VERSION : 0.1
BEGIN

REGION Network 1
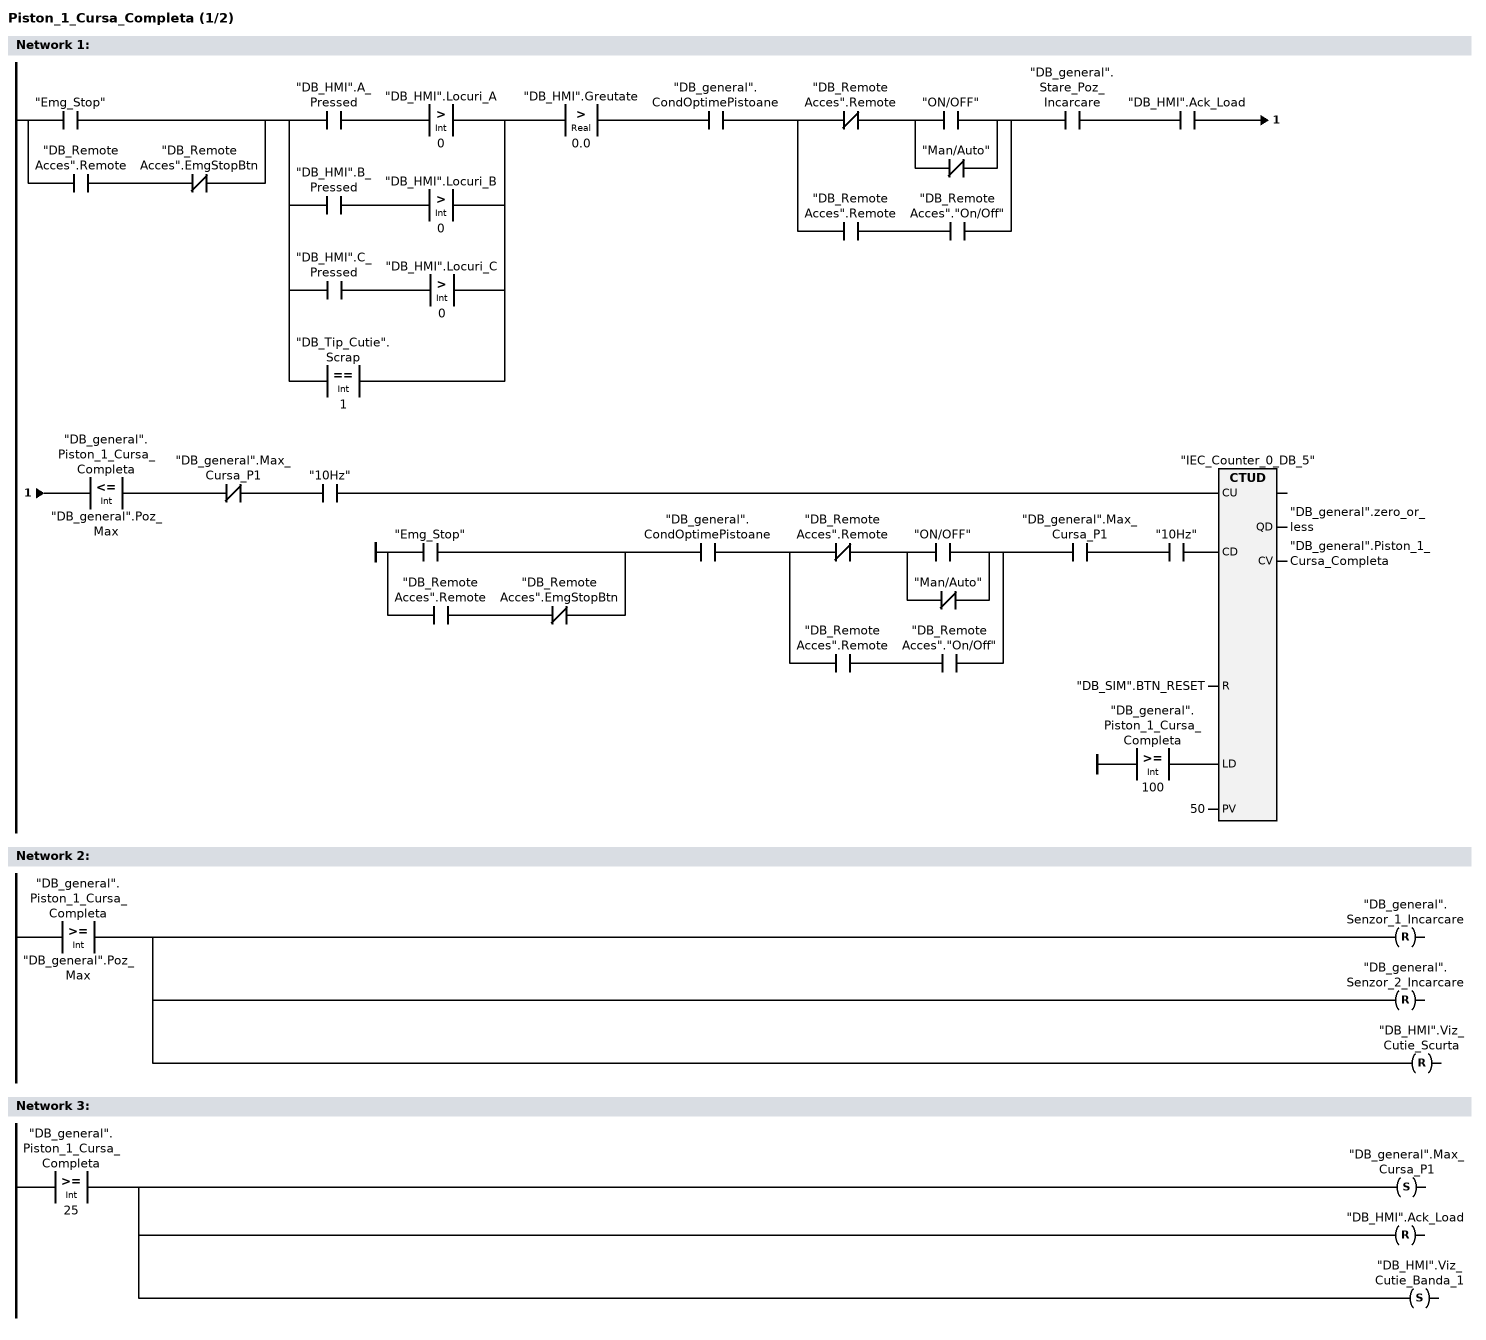
   "IEC_Counter_0_DB_5".CTUD(CU := ("Emg_Stop" OR ("DB_RemoteAcces".Remote AND NOT "DB_RemoteAcces".EmgStopBtn)) AND (("DB_HMI".A_Pressed AND ("DB_HMI".Locuri_A > 0)) OR ("DB_HMI".B_Pressed AND ("DB_HMI".Locuri_B > 0)) OR ("DB_HMI".C_Pressed AND ("DB_HMI".Locuri_C > 0)) OR ("DB_Tip_Cutie".Scrap = 1)) AND ("DB_HMI".Greutate > 0.0) AND "DB_general".CondOptimePistoane AND ((NOT "DB_RemoteAcces".Remote AND ("ON/OFF" OR NOT "Man/Auto")) OR ("DB_RemoteAcces".Remote AND "DB_RemoteAcces"."On/Off")) AND "DB_general".Stare_Poz_Incarcare AND "DB_HMI".Ack_Load AND ("DB_general".Piston_1_Cursa_Completa <= "DB_general".Poz_Max) AND NOT "DB_general".Max_Cursa_P1 AND "10Hz",
                           CD := ("Emg_Stop" OR ("DB_RemoteAcces".Remote AND NOT "DB_RemoteAcces".EmgStopBtn)) AND "DB_general".CondOptimePistoane AND ((NOT "DB_RemoteAcces".Remote AND ("ON/OFF" OR NOT "Man/Auto")) OR ("DB_RemoteAcces".Remote AND "DB_RemoteAcces"."On/Off")) AND "DB_general".Max_Cursa_P1 AND "10Hz",
                           R := "DB_SIM".BTN_RESET,
                           LD := "DB_general".Piston_1_Cursa_Completa >= 100,
                           PV := 50,
                           QD => "DB_general".zero_or_less,
                           CV => "DB_general".Piston_1_Cursa_Completa);
END_REGION

REGION Network 2
   RUNG wire#powerrail
      { S7_Templates := "SrcType := Int" } GE_Contact(in1 := "DB_general".Piston_1_Cursa_Completa, in2 := "DB_general".Poz_Max)
      wire#w1
      R_Coil( "DB_general".Senzor_1_Incarcare )
   END_RUNG
   RUNG wire#w1
      R_Coil( "DB_general".Senzor_2_Incarcare )
   END_RUNG
   RUNG wire#w1
      R_Coil( "DB_HMI".Viz_Cutie_Scurta )
   END_RUNG
   // the same network as SCL:
   IF "DB_general".Piston_1_Cursa_Completa >= "DB_general".Poz_Max THEN
       "DB_general".Senzor_1_Incarcare := FALSE;
       "DB_general".Senzor_2_Incarcare := FALSE;
       "DB_HMI".Viz_Cutie_Scurta := FALSE;
   END_IF;
END_REGION

REGION Network 3
   RUNG wire#powerrail
      { S7_Templates := "SrcType := Int" } GE_Contact(in1 := "DB_general".Piston_1_Cursa_Completa, in2 := 25)
      wire#w1
      S_Coil( "DB_general".Max_Cursa_P1 )
   END_RUNG
   RUNG wire#w1
      R_Coil( "DB_HMI".Ack_Load )
   END_RUNG
   RUNG wire#w1
      S_Coil( "DB_HMI".Viz_Cutie_Banda_1 )
   END_RUNG
   // the same network as SCL:
   IF "DB_general".Piston_1_Cursa_Completa >= 25 THEN
       "DB_general".Max_Cursa_P1 := TRUE;
       "DB_HMI".Ack_Load := FALSE;
       "DB_HMI".Viz_Cutie_Banda_1 := TRUE;
   END_IF;
END_REGION

REGION Network 4
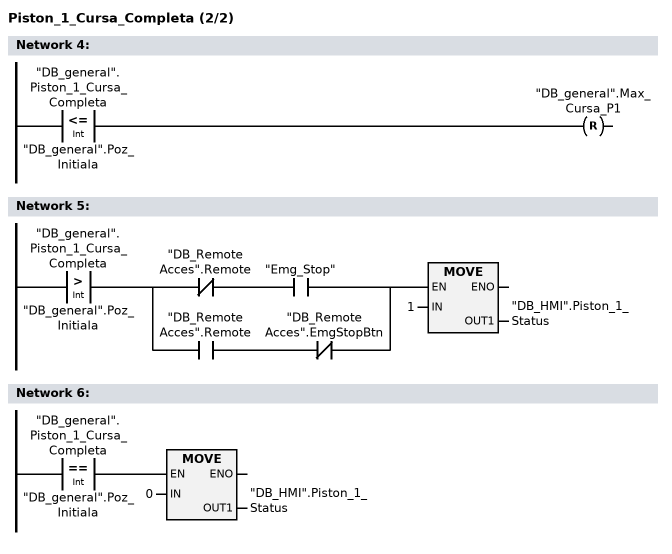
   RUNG wire#powerrail
      { S7_Templates := "SrcType := Int" } LE_Contact(in1 := "DB_general".Piston_1_Cursa_Completa, in2 := "DB_general".Poz_Initiala)
      R_Coil( "DB_general".Max_Cursa_P1 )
   END_RUNG
   // the same network as SCL:
   IF "DB_general".Piston_1_Cursa_Completa <= "DB_general".Poz_Initiala THEN
       "DB_general".Max_Cursa_P1 := FALSE;
   END_IF;
END_REGION

REGION Network 5
   RUNG wire#powerrail
      { S7_Templates := "SrcType := Int" } GT_Contact(in1 := "DB_general".Piston_1_Cursa_Completa, in2 := "DB_general".Poz_Initiala)
      wire#w1
      I_Contact( "DB_RemoteAcces".Remote )
      Contact( "Emg_Stop" )
      wire#w2
      { S7_GenerateENO := "TRUE" } Move(in := 1, out1 => "DB_HMI".Piston_1_Status)
   END_RUNG
   RUNG wire#w1
      Contact( "DB_RemoteAcces".Remote )
      I_Contact( "DB_RemoteAcces".EmgStopBtn )
   END_RUNG wire#w2
   // the same network as SCL:
   IF ("DB_general".Piston_1_Cursa_Completa > "DB_general".Poz_Initiala) AND ((NOT "DB_RemoteAcces".Remote AND "Emg_Stop") OR ("DB_RemoteAcces".Remote AND NOT "DB_RemoteAcces".EmgStopBtn)) THEN
       "DB_HMI".Piston_1_Status := 1;
   END_IF;
END_REGION

REGION Network 6
   RUNG wire#powerrail
      { S7_Templates := "SrcType := Int" } EQ_Contact(in1 := "DB_general".Piston_1_Cursa_Completa, in2 := "DB_general".Poz_Initiala)
      { S7_GenerateENO := "TRUE" } Move(in := 0, out1 => "DB_HMI".Piston_1_Status)
   END_RUNG
   // the same network as SCL:
   IF "DB_general".Piston_1_Cursa_Completa = "DB_general".Poz_Initiala THEN
       "DB_HMI".Piston_1_Status := 0;
   END_IF;
END_REGION
END_FUNCTION_BLOCK

FUNCTION_BLOCK "Piston_2_Cursa_Completa"   // FB17, LAD
{ S7_Optimized_Access := 'FALSE' }
VERSION : 0.1
BEGIN

REGION Network 1
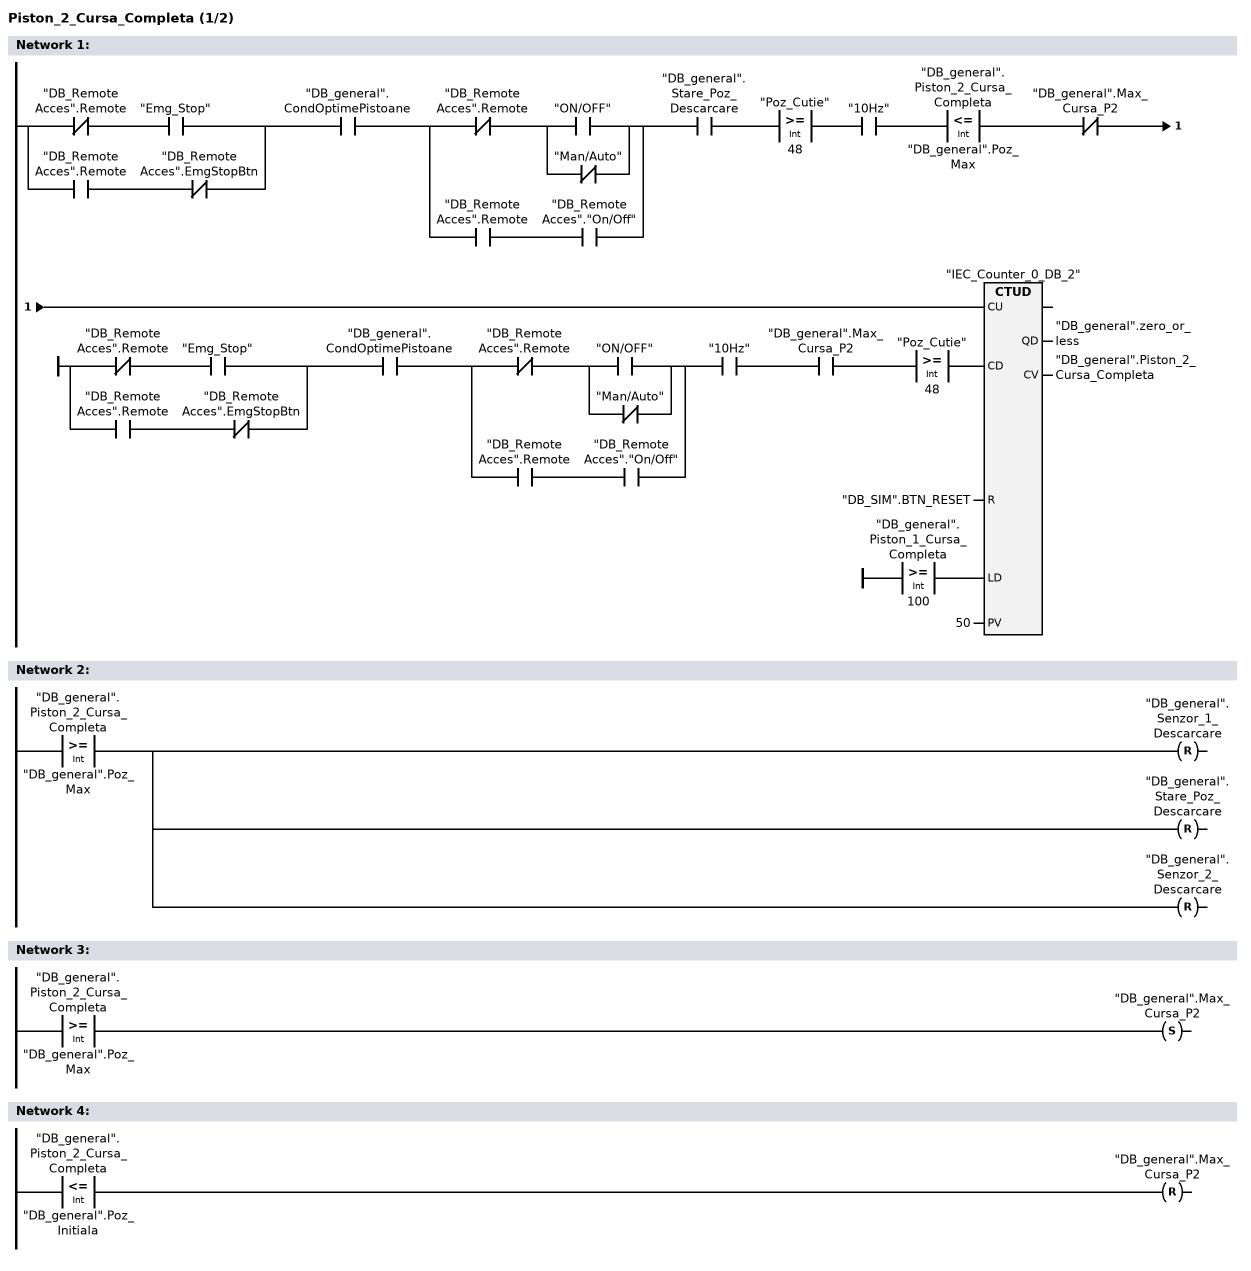
   "IEC_Counter_0_DB_2".CTUD(CU := ((NOT "DB_RemoteAcces".Remote AND "Emg_Stop") OR ("DB_RemoteAcces".Remote AND NOT "DB_RemoteAcces".EmgStopBtn)) AND "DB_general".CondOptimePistoane AND ((NOT "DB_RemoteAcces".Remote AND ("ON/OFF" OR NOT "Man/Auto")) OR ("DB_RemoteAcces".Remote AND "DB_RemoteAcces"."On/Off")) AND "DB_general".Stare_Poz_Descarcare AND ("Poz_Cutie" >= 48) AND "10Hz" AND ("DB_general".Piston_2_Cursa_Completa <= "DB_general".Poz_Max) AND NOT "DB_general".Max_Cursa_P2,
                           CD := ((NOT "DB_RemoteAcces".Remote AND "Emg_Stop") OR ("DB_RemoteAcces".Remote AND NOT "DB_RemoteAcces".EmgStopBtn)) AND "DB_general".CondOptimePistoane AND ((NOT "DB_RemoteAcces".Remote AND ("ON/OFF" OR NOT "Man/Auto")) OR ("DB_RemoteAcces".Remote AND "DB_RemoteAcces"."On/Off")) AND "10Hz" AND "DB_general".Max_Cursa_P2 AND ("Poz_Cutie" >= 48),
                           R := "DB_SIM".BTN_RESET,
                           LD := "DB_general".Piston_1_Cursa_Completa >= 100,
                           PV := 50,
                           QD => "DB_general".zero_or_less,
                           CV => "DB_general".Piston_2_Cursa_Completa);
END_REGION

REGION Network 2
   RUNG wire#powerrail
      { S7_Templates := "SrcType := Int" } GE_Contact(in1 := "DB_general".Piston_2_Cursa_Completa, in2 := "DB_general".Poz_Max)
      wire#w1
      R_Coil( "DB_general".Senzor_1_Descarcare )
   END_RUNG
   RUNG wire#w1
      R_Coil( "DB_general".Stare_Poz_Descarcare )
   END_RUNG
   RUNG wire#w1
      R_Coil( "DB_general".Senzor_2_Descarcare )
   END_RUNG
   // the same network as SCL:
   IF "DB_general".Piston_2_Cursa_Completa >= "DB_general".Poz_Max THEN
       "DB_general".Senzor_1_Descarcare := FALSE;
       "DB_general".Stare_Poz_Descarcare := FALSE;
       "DB_general".Senzor_2_Descarcare := FALSE;
   END_IF;
END_REGION

REGION Network 3
   RUNG wire#powerrail
      { S7_Templates := "SrcType := Int" } GE_Contact(in1 := "DB_general".Piston_2_Cursa_Completa, in2 := "DB_general".Poz_Max)
      S_Coil( "DB_general".Max_Cursa_P2 )
   END_RUNG
   // the same network as SCL:
   IF "DB_general".Piston_2_Cursa_Completa >= "DB_general".Poz_Max THEN
       "DB_general".Max_Cursa_P2 := TRUE;
   END_IF;
END_REGION

REGION Network 4
   RUNG wire#powerrail
      { S7_Templates := "SrcType := Int" } LE_Contact(in1 := "DB_general".Piston_2_Cursa_Completa, in2 := "DB_general".Poz_Initiala)
      R_Coil( "DB_general".Max_Cursa_P2 )
   END_RUNG
   // the same network as SCL:
   IF "DB_general".Piston_2_Cursa_Completa <= "DB_general".Poz_Initiala THEN
       "DB_general".Max_Cursa_P2 := FALSE;
   END_IF;
END_REGION

REGION Network 5
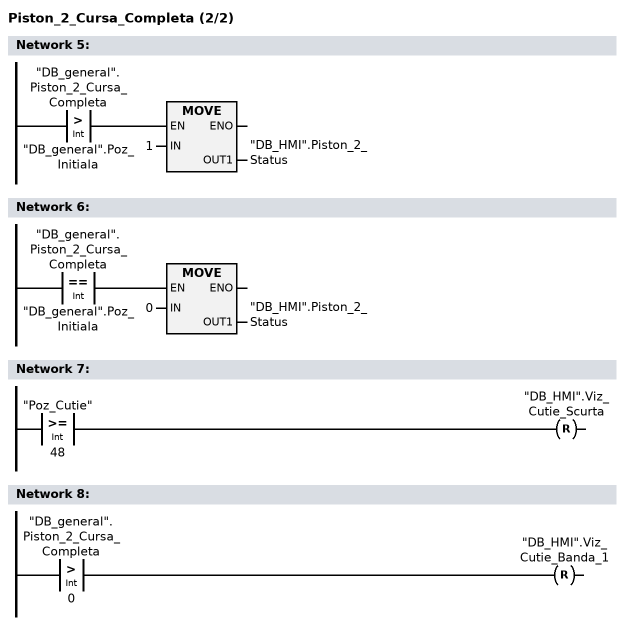
   RUNG wire#powerrail
      { S7_Templates := "SrcType := Int" } GT_Contact(in1 := "DB_general".Piston_2_Cursa_Completa, in2 := "DB_general".Poz_Initiala)
      { S7_GenerateENO := "TRUE" } Move(in := 1, out1 => "DB_HMI".Piston_2_Status)
   END_RUNG
   // the same network as SCL:
   IF "DB_general".Piston_2_Cursa_Completa > "DB_general".Poz_Initiala THEN
       "DB_HMI".Piston_2_Status := 1;
   END_IF;
END_REGION

REGION Network 6
   RUNG wire#powerrail
      { S7_Templates := "SrcType := Int" } EQ_Contact(in1 := "DB_general".Piston_2_Cursa_Completa, in2 := "DB_general".Poz_Initiala)
      { S7_GenerateENO := "TRUE" } Move(in := 0, out1 => "DB_HMI".Piston_2_Status)
   END_RUNG
   // the same network as SCL:
   IF "DB_general".Piston_2_Cursa_Completa = "DB_general".Poz_Initiala THEN
       "DB_HMI".Piston_2_Status := 0;
   END_IF;
END_REGION

REGION Network 7
   RUNG wire#powerrail
      { S7_Templates := "SrcType := Int" } GE_Contact(in1 := "Poz_Cutie", in2 := 48)
      R_Coil( "DB_HMI".Viz_Cutie_Scurta )
   END_RUNG
   // the same network as SCL:
   IF "Poz_Cutie" >= 48 THEN "DB_HMI".Viz_Cutie_Scurta := FALSE; END_IF;
END_REGION

REGION Network 8
   RUNG wire#powerrail
      { S7_Templates := "SrcType := Int" } GT_Contact(in1 := "DB_general".Piston_2_Cursa_Completa, in2 := 0)
      R_Coil( "DB_HMI".Viz_Cutie_Banda_1 )
   END_RUNG
   // the same network as SCL:
   IF "DB_general".Piston_2_Cursa_Completa > 0 THEN "DB_HMI".Viz_Cutie_Banda_1 := FALSE; END_IF;
END_REGION
END_FUNCTION_BLOCK

// folder: Statie Distribuire/Functii

FUNCTION_BLOCK "Banda_1"   // FB4, SCL
{ S7_Optimized_Access := 'FALSE' }
VERSION : 0.1
   VAR_INPUT
      Stare_Poz_Incarcare : Bool;
      Stare_Poz_Descarcare : Bool;
      Stare_Descarcare : Bool;   // Acesta este o valoare de test in care urm ca la finalul de cursa (Animatie Banda 1) pozitia descarcare sa fie facuta adev
      "Man/Auto" : Bool;
      Btn_LOAD : Bool;
   END_VAR
   VAR_OUTPUT
      Status_Banda_1 : Bool;
   END_VAR
   VAR
      Status_Poz_Cantar : Bool;
      Greutate_cantar : Int;
      Limitare_Interval : Bool;
      "ON/OFF" : Bool;
      Start_Pressed : Bool;
      AFost : Bool;
      Aux : Bool;
      LOAD_Pressed : Bool;
   END_VAR
BEGIN
   //MOD MANUAL/AUTOMAT + BUTOANE MANUAL
   IF #"Man/Auto"  THEN//daca e modul manual poti actiona butoane  true e manual false e automat

       IF "Start"  THEN
           #"Start_Pressed" := TRUE;  // setare variabila aux
           #"ON/OFF" := #Start_Pressed;
           "ON/OFF" := #"ON/OFF";
       END_IF;

       IF  "Stop"=TRUE  THEN
           #"ON/OFF" := #Start_Pressed;  //atribuire var aux
           "ON/OFF" := #"ON/OFF";
       ELSE
           IF "Stop" = FALSE THEN
               #"ON/OFF" := FALSE;
               "ON/OFF" := #"ON/OFF";
               #"Start_Pressed" := FALSE;
           END_IF;// reset variabila auxiliară la apasare stop
       END_IF;
       IF "Emg_Stop" = TRUE  THEN
           #"ON/OFF" := #Start_Pressed;  //atribuire var aux
       ELSE
           IF "Emg_Stop" = FALSE  THEN
               #"ON/OFF" := FALSE;
               "ON/OFF" := #"ON/OFF";
               #"Start_Pressed" := FALSE;
           END_IF;// reset variabila auxiliară la apasare stop
       END_IF;


   ELSE
      // #"ON/OFF" := FALSE;
      // "ON/OFF" := #"ON/OFF";
      #"Start_Pressed" := FALSE;  // Resetați variabila auxiliară în modul Manual


   END_IF;


   //LIMITARI CAPAT DE BANDA

   IF #Stare_Poz_Incarcare AND #Stare_Poz_Descarcare = FALSE AND #Stare_Descarcare=FALSE THEN//limitari de la sezorii din capetele benzii
       #Limitare_Interval := FALSE; //daca e prezent la primul nu porneste 
   ELSE
       IF #Stare_Poz_Incarcare = FALSE AND #Stare_Poz_Descarcare AND #Stare_Descarcare THEN
         #Limitare_Interval := FALSE;//daca e prezent la al doilea se opreste banda
     ELSE
         #Limitare_Interval := TRUE;

     END_IF;


   END_IF;
   // Logica pentru setare și resetare


   //START MOTOARE 
   IF #Btn_LOAD THEN
       #LOAD_Pressed := true;
   END_IF;

   IF "Poz_Cutie"<=100 THEN

       #LOAD_Pressed := TRUE;

   ELSE
       #LOAD_Pressed := FALSE;
       // Statement section IF
       ;
   END_IF;

   IF "DB_RemoteAcces"."Remote" = FALSE THEN

       IF "Man/Auto" THEN
           IF "Emg_Stop" = TRUE AND #"ON/OFF" = TRUE AND #Limitare_Interval AND "DB_HMI".BTN_LOAD THEN


               #Status_Banda_1 := TRUE;

           ELSE

               #Status_Banda_1 := FALSE;
           END_IF;

       ELSE
           IF "Emg_Stop" = TRUE AND #Limitare_Interval AND "DB_HMI".BTN_LOAD THEN

               #Status_Banda_1 := TRUE;
           ELSE

               #Status_Banda_1 := FALSE;
           END_IF;


       END_IF;


   ELSE
       IF "DB_RemoteAcces"."Remote" = TRUE THEN
           IF "DB_RemoteAcces"."Manual/Auto" = FALSE THEN
               IF "DB_RemoteAcces".EmgStopBtn = FALSE AND "DB_RemoteAcces"."On/Off" = TRUE AND #Limitare_Interval AND "DB_HMI".BTN_LOAD THEN


                   #Status_Banda_1 := TRUE;

               ELSE

                   #Status_Banda_1 := FALSE;
               END_IF;

           ELSE
               IF "DB_RemoteAcces".EmgStopBtn= FALSE AND "DB_RemoteAcces"."On/Off" = TRUE AND #Limitare_Interval AND"DB_HMI".BTN_LOAD THEN

                   #Status_Banda_1 := TRUE;
               ELSE

                   #Status_Banda_1 := FALSE;
               END_IF;


           END_IF;
       END_IF;

   END_IF;
END_FUNCTION_BLOCK

FUNCTION_BLOCK "Cantar"   // FB6, SCL
{ S7_Optimized_Access := 'FALSE' }
VERSION : 0.1
   VAR_INPUT
      Status_Poz : Bool;
      emgy_ok : Bool;
   END_VAR
   VAR_OUTPUT
      Greutate : Int;
   END_VAR
   VAR
      time_struct : Struct
         an : Byte;
         luna : Byte;
         zi : Byte;
         ora : Byte;
         minut : Byte;
         sec : Byte;
         milisec : Byte;
         weekday : Byte;
      END_STRUCT;
      rand : Int;
      i : Int;
      val : Int := 100;
   END_VAR
BEGIN

   #val := 100;

   IF "Emg_Stop" = TRUE THEN

       IF #Status_Poz = TRUE THEN

           FOR #i := 0 TO 9 DO
               #val := #val + 5;
               #Greutate := #val;
               END_FOR;


       END_IF;

   END_IF;
END_FUNCTION_BLOCK

FUNCTION_BLOCK "Verificare_Poz_StartSec"   // FB7, SCL
{ S7_Optimized_Access := 'FALSE' }
VERSION : 0.1
   VAR_INPUT
      Senzor_1 : Bool;
      Senzor_2 : Bool;
   END_VAR
   VAR_OUTPUT
      Status_Poz : Bool := false;
   END_VAR
BEGIN


       IF #Senzor_1 = TRUE AND #Senzor_2 = TRUE THEN
           #Status_Poz := TRUE;  // verif pozitie
       ELSE
           #Status_Poz := FALSE;
       END_IF;
END_FUNCTION_BLOCK

FUNCTION "Control_Enable" : Void   // FC12, LAD
{ S7_Optimized_Access := 'FALSE' }
VERSION : 0.1
BEGIN

REGION Network 1: Btn de load / Schaltfläche „Laden“
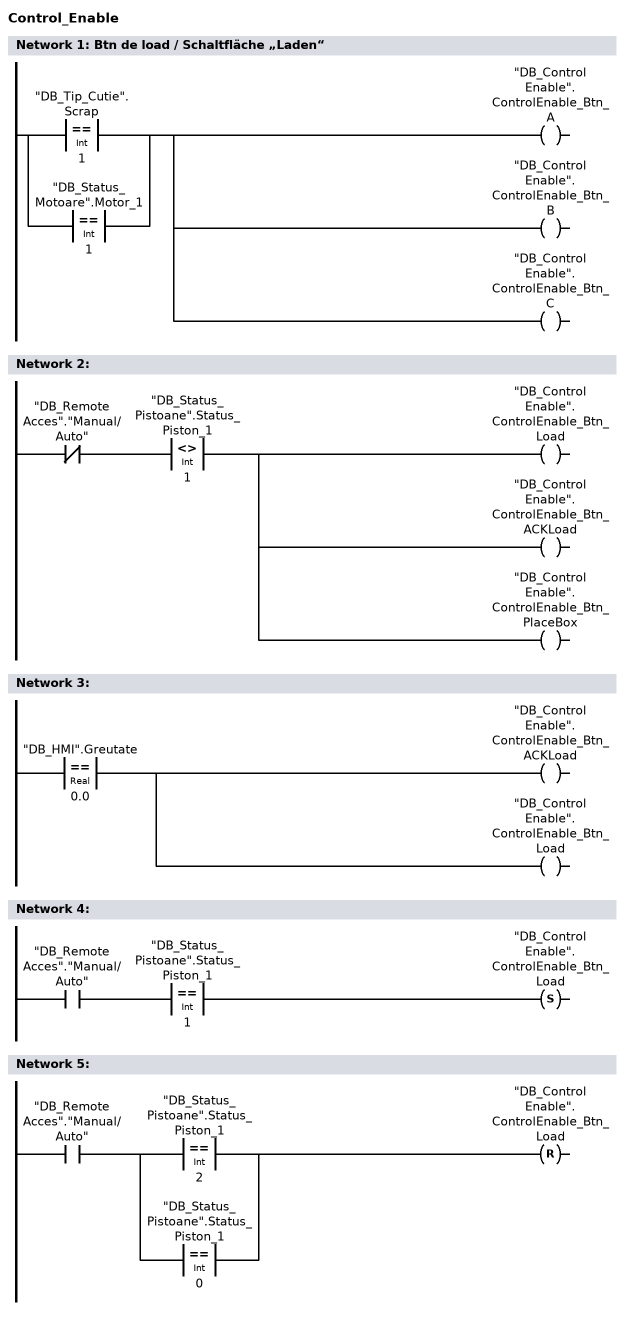
   RUNG wire#powerrail
      { S7_Templates := "SrcType := Int" } EQ_Contact(in1 := "DB_Tip_Cutie".Scrap, in2 := 1)
      wire#w1
      Coil( "DB_ControlEnable".ControlEnable_Btn_A )
   END_RUNG
   RUNG wire#powerrail
      { S7_Templates := "SrcType := Int" } EQ_Contact(in1 := "DB_Status_Motoare".Motor_1, in2 := 1)
   END_RUNG wire#w1
   RUNG wire#w1
      Coil( "DB_ControlEnable".ControlEnable_Btn_B )
   END_RUNG
   RUNG wire#w1
      Coil( "DB_ControlEnable".ControlEnable_Btn_C )
   END_RUNG
   // the same network as SCL:
   "DB_ControlEnable".ControlEnable_Btn_A := ("DB_Tip_Cutie".Scrap = 1) OR ("DB_Status_Motoare".Motor_1 = 1);
   "DB_ControlEnable".ControlEnable_Btn_B := "DB_ControlEnable".ControlEnable_Btn_A;
   "DB_ControlEnable".ControlEnable_Btn_C := "DB_ControlEnable".ControlEnable_Btn_A;
END_REGION

REGION Network 2
   RUNG wire#powerrail
      I_Contact( "DB_RemoteAcces"."Manual/Auto" )
      { S7_Templates := "SrcType := Int" } NE_Contact(in1 := "DB_Status_Pistoane".Status_Piston_1, in2 := 1)
      wire#w1
      Coil( "DB_ControlEnable".ControlEnable_Btn_Load )
   END_RUNG
   RUNG wire#w1
      Coil( "DB_ControlEnable".ControlEnable_Btn_ACKLoad )
   END_RUNG
   RUNG wire#w1
      Coil( "DB_ControlEnable".ControlEnable_Btn_PlaceBox )
   END_RUNG
   // the same network as SCL:
   "DB_ControlEnable".ControlEnable_Btn_Load := NOT "DB_RemoteAcces"."Manual/Auto" AND ("DB_Status_Pistoane".Status_Piston_1 <> 1);
   "DB_ControlEnable".ControlEnable_Btn_ACKLoad := "DB_ControlEnable".ControlEnable_Btn_Load;
   "DB_ControlEnable".ControlEnable_Btn_PlaceBox := "DB_ControlEnable".ControlEnable_Btn_Load;
END_REGION

REGION Network 3
   RUNG wire#powerrail
      { S7_Templates := "SrcType := Real" } EQ_Contact(in1 := "DB_HMI".Greutate, in2 := 0.0)
      wire#w1
      Coil( "DB_ControlEnable".ControlEnable_Btn_ACKLoad )
   END_RUNG
   RUNG wire#w1
      Coil( "DB_ControlEnable".ControlEnable_Btn_Load )
   END_RUNG
   // the same network as SCL:
   "DB_ControlEnable".ControlEnable_Btn_ACKLoad := "DB_HMI".Greutate = 0.0;
   "DB_ControlEnable".ControlEnable_Btn_Load := "DB_ControlEnable".ControlEnable_Btn_ACKLoad;
END_REGION

REGION Network 4
   RUNG wire#powerrail
      Contact( "DB_RemoteAcces"."Manual/Auto" )
      { S7_Templates := "SrcType := Int" } EQ_Contact(in1 := "DB_Status_Pistoane".Status_Piston_1, in2 := 1)
      S_Coil( "DB_ControlEnable".ControlEnable_Btn_Load )
   END_RUNG
   // the same network as SCL:
   IF "DB_RemoteAcces"."Manual/Auto" AND ("DB_Status_Pistoane".Status_Piston_1 = 1) THEN
       "DB_ControlEnable".ControlEnable_Btn_Load := TRUE;
   END_IF;
END_REGION

REGION Network 5
   RUNG wire#powerrail
      Contact( "DB_RemoteAcces"."Manual/Auto" )
      wire#w1
      { S7_Templates := "SrcType := Int" } EQ_Contact(in1 := "DB_Status_Pistoane".Status_Piston_1, in2 := 2)
      wire#w2
      R_Coil( "DB_ControlEnable".ControlEnable_Btn_Load )
   END_RUNG
   RUNG wire#w1
      { S7_Templates := "SrcType := Int" } EQ_Contact(in1 := "DB_Status_Pistoane".Status_Piston_1, in2 := 0)
   END_RUNG wire#w2
   // the same network as SCL:
   IF "DB_RemoteAcces"."Manual/Auto" AND (("DB_Status_Pistoane".Status_Piston_1 = 2) OR ("DB_Status_Pistoane".Status_Piston_1 = 0)) THEN
       "DB_ControlEnable".ControlEnable_Btn_Load := FALSE;
   END_IF;
END_REGION
END_FUNCTION

FUNCTION "StatusBtnDistribuire" : Void   // FC13, LAD
{ S7_Optimized_Access := 'FALSE' }
VERSION : 0.1
BEGIN

REGION Network 1
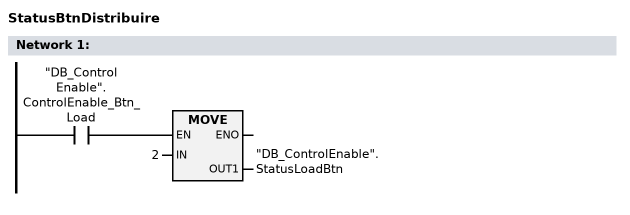
   RUNG wire#powerrail
      Contact( "DB_ControlEnable".ControlEnable_Btn_Load )
      { S7_GenerateENO := "TRUE" } Move(in := 2, out1 => "DB_ControlEnable".StatusLoadBtn)
   END_RUNG
   // the same network as SCL:
   IF "DB_ControlEnable".ControlEnable_Btn_Load THEN "DB_ControlEnable".StatusLoadBtn := 2; END_IF;
END_REGION
END_FUNCTION

// folder: Statie Incarcare/Animatii

FUNCTION_BLOCK "Animatie_Banda_Bile"   // FB15, LAD
{ S7_Optimized_Access := 'FALSE' }
VERSION : 0.1
   VAR_INPUT
      Status_Banda_2 : Bool;
      Btn_Transport : Bool;
   END_VAR
BEGIN

REGION Network 1
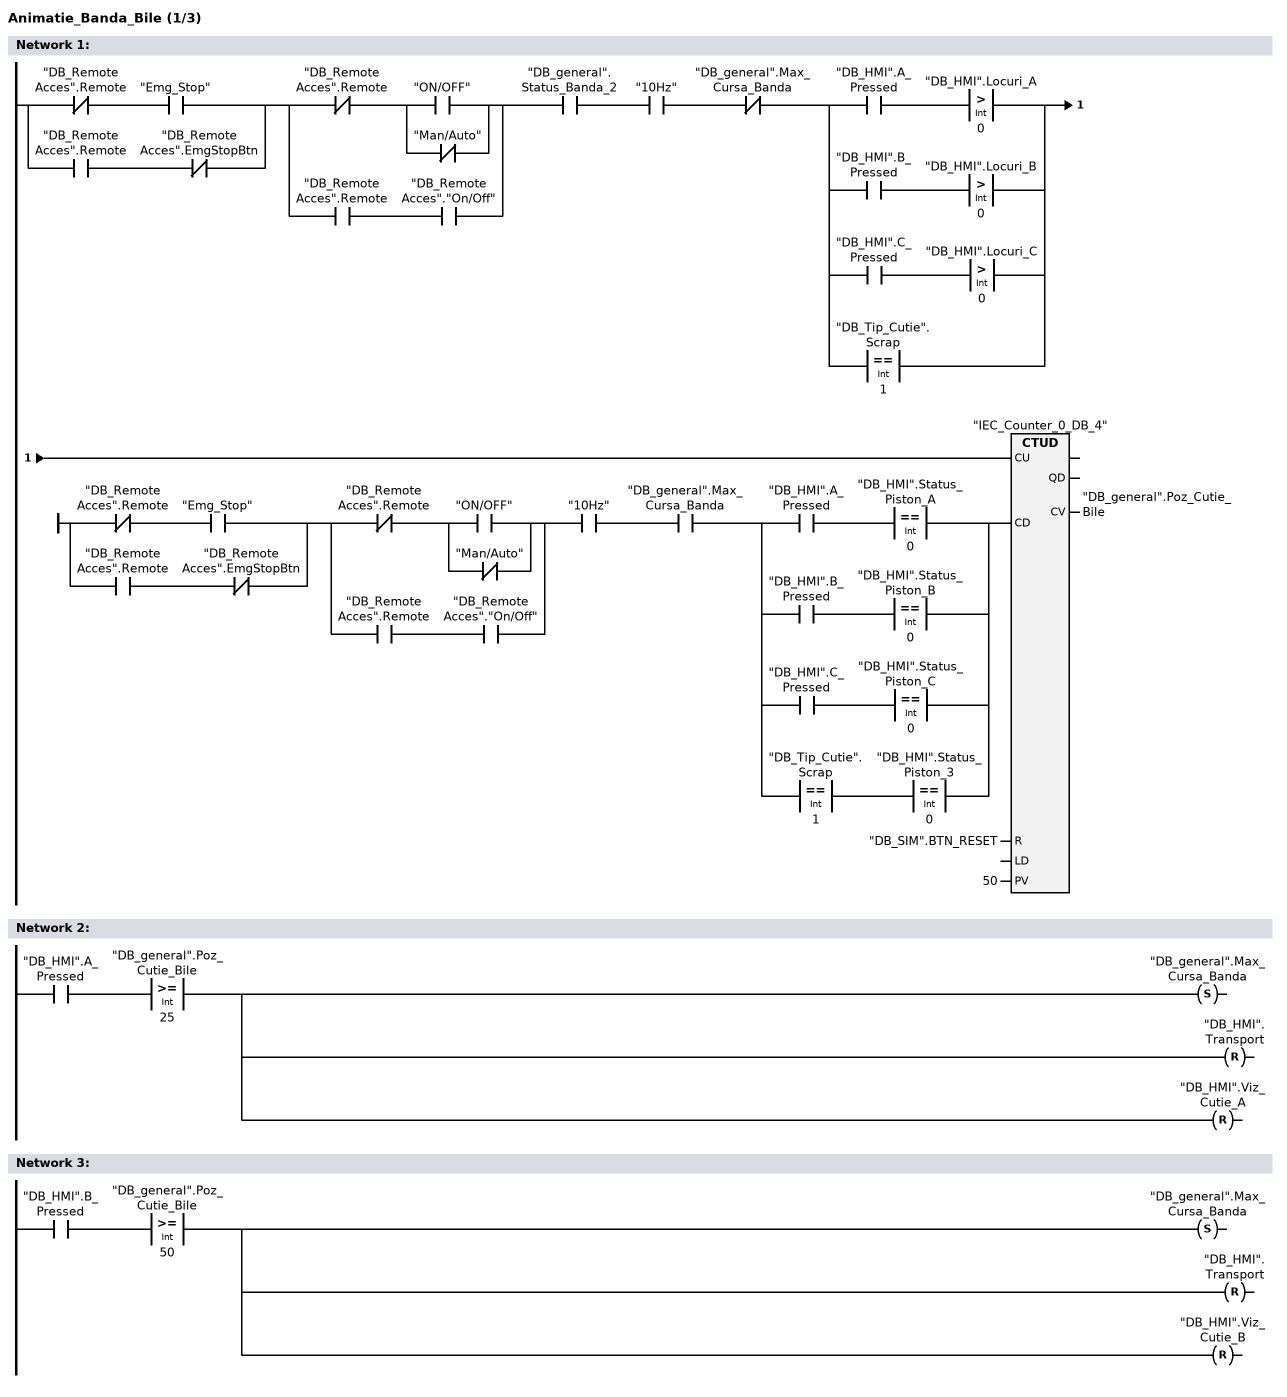
   "IEC_Counter_0_DB_4".CTUD(CU := ((NOT "DB_RemoteAcces".Remote AND "Emg_Stop") OR ("DB_RemoteAcces".Remote AND NOT "DB_RemoteAcces".EmgStopBtn)) AND ((NOT "DB_RemoteAcces".Remote AND ("ON/OFF" OR NOT "Man/Auto")) OR ("DB_RemoteAcces".Remote AND "DB_RemoteAcces"."On/Off")) AND "DB_general".Status_Banda_2 AND "10Hz" AND NOT "DB_general".Max_Cursa_Banda AND (("DB_HMI".A_Pressed AND ("DB_HMI".Locuri_A > 0)) OR ("DB_HMI".B_Pressed AND ("DB_HMI".Locuri_B > 0)) OR ("DB_HMI".C_Pressed AND ("DB_HMI".Locuri_C > 0)) OR ("DB_Tip_Cutie".Scrap = 1)),
                           CD := ((NOT "DB_RemoteAcces".Remote AND "Emg_Stop") OR ("DB_RemoteAcces".Remote AND NOT "DB_RemoteAcces".EmgStopBtn)) AND ((NOT "DB_RemoteAcces".Remote AND ("ON/OFF" OR NOT "Man/Auto")) OR ("DB_RemoteAcces".Remote AND "DB_RemoteAcces"."On/Off")) AND "10Hz" AND "DB_general".Max_Cursa_Banda AND (("DB_HMI".A_Pressed AND ("DB_HMI".Status_Piston_A = 0)) OR ("DB_HMI".B_Pressed AND ("DB_HMI".Status_Piston_B = 0)) OR ("DB_HMI".C_Pressed AND ("DB_HMI".Status_Piston_C = 0)) OR (("DB_Tip_Cutie".Scrap = 1) AND ("DB_HMI".Status_Piston_3 = 0))),
                           R := "DB_SIM".BTN_RESET,
                           PV := 50,
                           CV => "DB_general".Poz_Cutie_Bile);
END_REGION

REGION Network 2
   RUNG wire#powerrail
      Contact( "DB_HMI".A_Pressed )
      { S7_Templates := "SrcType := Int" } GE_Contact(in1 := "DB_general".Poz_Cutie_Bile, in2 := 25)
      wire#w1
      S_Coil( "DB_general".Max_Cursa_Banda )
   END_RUNG
   RUNG wire#w1
      R_Coil( "DB_HMI".Transport )
   END_RUNG
   RUNG wire#w1
      R_Coil( "DB_HMI".Viz_Cutie_A )
   END_RUNG
   // the same network as SCL:
   IF "DB_HMI".A_Pressed AND ("DB_general".Poz_Cutie_Bile >= 25) THEN
       "DB_general".Max_Cursa_Banda := TRUE;
       "DB_HMI".Transport := FALSE;
       "DB_HMI".Viz_Cutie_A := FALSE;
   END_IF;
END_REGION

REGION Network 3
   RUNG wire#powerrail
      Contact( "DB_HMI".B_Pressed )
      { S7_Templates := "SrcType := Int" } GE_Contact(in1 := "DB_general".Poz_Cutie_Bile, in2 := 50)
      wire#w1
      S_Coil( "DB_general".Max_Cursa_Banda )
   END_RUNG
   RUNG wire#w1
      R_Coil( "DB_HMI".Transport )
   END_RUNG
   RUNG wire#w1
      R_Coil( "DB_HMI".Viz_Cutie_B )
   END_RUNG
   // the same network as SCL:
   IF "DB_HMI".B_Pressed AND ("DB_general".Poz_Cutie_Bile >= 50) THEN
       "DB_general".Max_Cursa_Banda := TRUE;
       "DB_HMI".Transport := FALSE;
       "DB_HMI".Viz_Cutie_B := FALSE;
   END_IF;
END_REGION

REGION Network 4
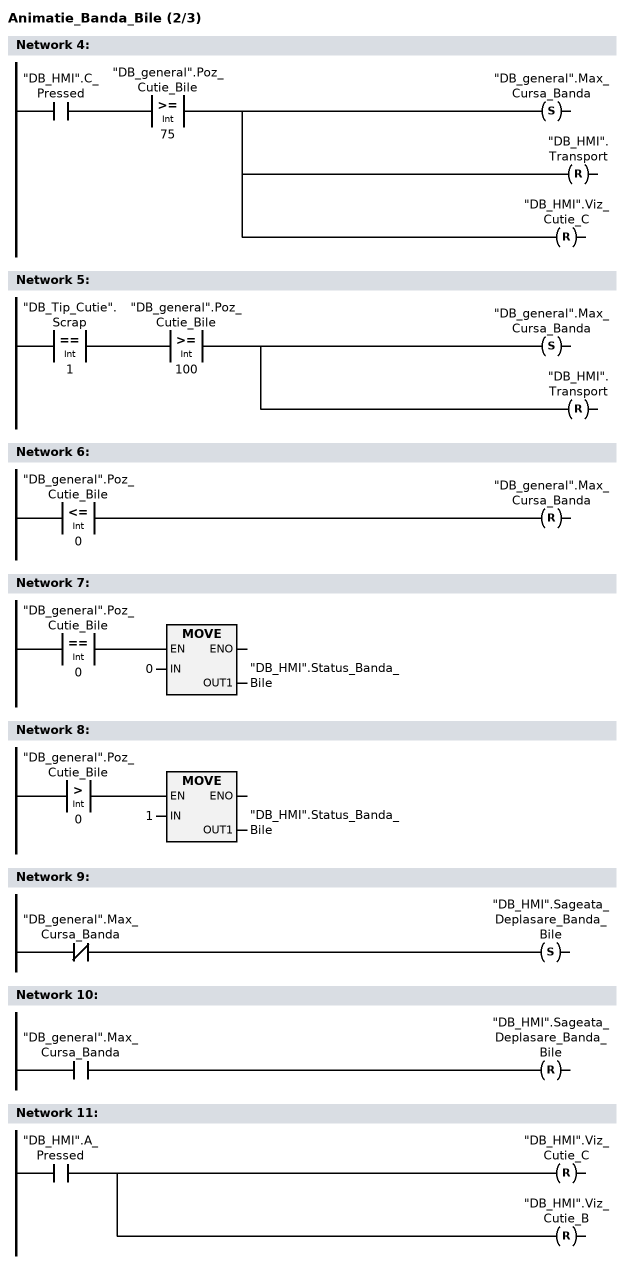
   RUNG wire#powerrail
      Contact( "DB_HMI".C_Pressed )
      { S7_Templates := "SrcType := Int" } GE_Contact(in1 := "DB_general".Poz_Cutie_Bile, in2 := 75)
      wire#w1
      S_Coil( "DB_general".Max_Cursa_Banda )
   END_RUNG
   RUNG wire#w1
      R_Coil( "DB_HMI".Transport )
   END_RUNG
   RUNG wire#w1
      R_Coil( "DB_HMI".Viz_Cutie_C )
   END_RUNG
   // the same network as SCL:
   IF "DB_HMI".C_Pressed AND ("DB_general".Poz_Cutie_Bile >= 75) THEN
       "DB_general".Max_Cursa_Banda := TRUE;
       "DB_HMI".Transport := FALSE;
       "DB_HMI".Viz_Cutie_C := FALSE;
   END_IF;
END_REGION

REGION Network 5
   RUNG wire#powerrail
      { S7_Templates := "SrcType := Int" } EQ_Contact(in1 := "DB_Tip_Cutie".Scrap, in2 := 1)
      { S7_Templates := "SrcType := Int" } GE_Contact(in1 := "DB_general".Poz_Cutie_Bile, in2 := 100)
      wire#w1
      S_Coil( "DB_general".Max_Cursa_Banda )
   END_RUNG
   RUNG wire#w1
      R_Coil( "DB_HMI".Transport )
   END_RUNG
   // the same network as SCL:
   IF ("DB_Tip_Cutie".Scrap = 1) AND ("DB_general".Poz_Cutie_Bile >= 100) THEN
       "DB_general".Max_Cursa_Banda := TRUE;
       "DB_HMI".Transport := FALSE;
   END_IF;
END_REGION

REGION Network 6
   RUNG wire#powerrail
      { S7_Templates := "SrcType := Int" } LE_Contact(in1 := "DB_general".Poz_Cutie_Bile, in2 := 0)
      R_Coil( "DB_general".Max_Cursa_Banda )
   END_RUNG
   // the same network as SCL:
   IF "DB_general".Poz_Cutie_Bile <= 0 THEN "DB_general".Max_Cursa_Banda := FALSE; END_IF;
END_REGION

REGION Network 7
   RUNG wire#powerrail
      { S7_Templates := "SrcType := Int" } EQ_Contact(in1 := "DB_general".Poz_Cutie_Bile, in2 := 0)
      { S7_GenerateENO := "TRUE" } Move(in := 0, out1 => "DB_HMI".Status_Banda_Bile)
   END_RUNG
   // the same network as SCL:
   IF "DB_general".Poz_Cutie_Bile = 0 THEN "DB_HMI".Status_Banda_Bile := 0; END_IF;
END_REGION

REGION Network 8
   RUNG wire#powerrail
      { S7_Templates := "SrcType := Int" } GT_Contact(in1 := "DB_general".Poz_Cutie_Bile, in2 := 0)
      { S7_GenerateENO := "TRUE" } Move(in := 1, out1 => "DB_HMI".Status_Banda_Bile)
   END_RUNG
   // the same network as SCL:
   IF "DB_general".Poz_Cutie_Bile > 0 THEN "DB_HMI".Status_Banda_Bile := 1; END_IF;
END_REGION

REGION Network 9
   RUNG wire#powerrail
      I_Contact( "DB_general".Max_Cursa_Banda )
      S_Coil( "DB_HMI".Sageata_Deplasare_Banda_Bile )
   END_RUNG
   // the same network as SCL:
   IF NOT "DB_general".Max_Cursa_Banda THEN "DB_HMI".Sageata_Deplasare_Banda_Bile := TRUE; END_IF;
END_REGION

REGION Network 10
   RUNG wire#powerrail
      Contact( "DB_general".Max_Cursa_Banda )
      R_Coil( "DB_HMI".Sageata_Deplasare_Banda_Bile )
   END_RUNG
   // the same network as SCL:
   IF "DB_general".Max_Cursa_Banda THEN "DB_HMI".Sageata_Deplasare_Banda_Bile := FALSE; END_IF;
END_REGION

REGION Network 11
   RUNG wire#powerrail
      Contact( "DB_HMI".A_Pressed )
      wire#w1
      R_Coil( "DB_HMI".Viz_Cutie_C )
   END_RUNG
   RUNG wire#w1
      R_Coil( "DB_HMI".Viz_Cutie_B )
   END_RUNG
   // the same network as SCL:
   IF "DB_HMI".A_Pressed THEN
       "DB_HMI".Viz_Cutie_C := FALSE;
       "DB_HMI".Viz_Cutie_B := FALSE;
   END_IF;
END_REGION

REGION Network 12
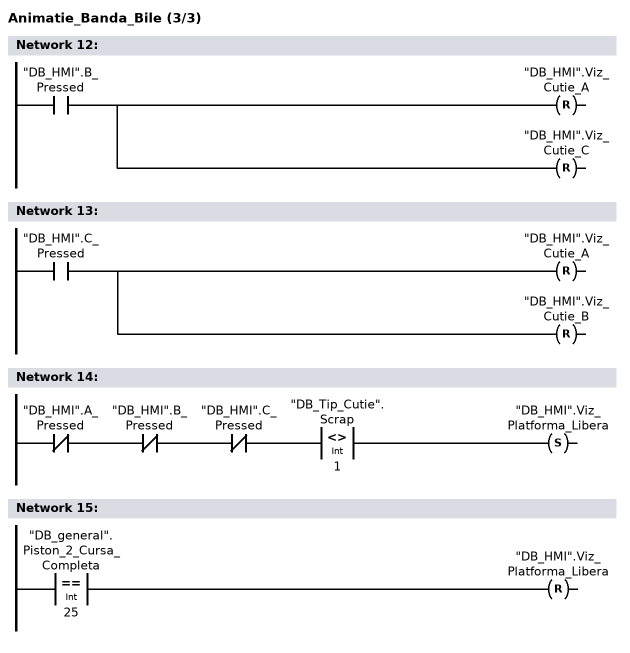
   RUNG wire#powerrail
      Contact( "DB_HMI".B_Pressed )
      wire#w1
      R_Coil( "DB_HMI".Viz_Cutie_A )
   END_RUNG
   RUNG wire#w1
      R_Coil( "DB_HMI".Viz_Cutie_C )
   END_RUNG
   // the same network as SCL:
   IF "DB_HMI".B_Pressed THEN
       "DB_HMI".Viz_Cutie_A := FALSE;
       "DB_HMI".Viz_Cutie_C := FALSE;
   END_IF;
END_REGION

REGION Network 13
   RUNG wire#powerrail
      Contact( "DB_HMI".C_Pressed )
      wire#w1
      R_Coil( "DB_HMI".Viz_Cutie_A )
   END_RUNG
   RUNG wire#w1
      R_Coil( "DB_HMI".Viz_Cutie_B )
   END_RUNG
   // the same network as SCL:
   IF "DB_HMI".C_Pressed THEN
       "DB_HMI".Viz_Cutie_A := FALSE;
       "DB_HMI".Viz_Cutie_B := FALSE;
   END_IF;
END_REGION

REGION Network 14
   RUNG wire#powerrail
      I_Contact( "DB_HMI".A_Pressed )
      I_Contact( "DB_HMI".B_Pressed )
      I_Contact( "DB_HMI".C_Pressed )
      { S7_Templates := "SrcType := Int" } NE_Contact(in1 := "DB_Tip_Cutie".Scrap, in2 := 1)
      S_Coil( "DB_HMI".Viz_Platforma_Libera )
   END_RUNG
   // the same network as SCL:
   IF NOT "DB_HMI".A_Pressed AND NOT "DB_HMI".B_Pressed AND NOT "DB_HMI".C_Pressed AND ("DB_Tip_Cutie".Scrap <> 1) THEN
       "DB_HMI".Viz_Platforma_Libera := TRUE;
   END_IF;
END_REGION
